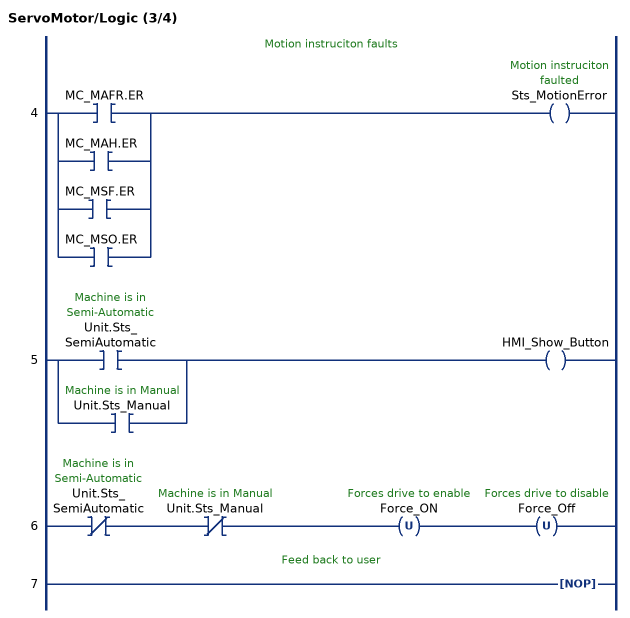
   // Motion instruciton faults
   4: [XIC(MC_MAFR.ER) ,XIC(MC_MAH.ER) ,XIC(MC_MSF.ER) ,XIC(MC_MSO.ER) ]OTE(Sts_MotionError);
   5: [XIC(Unit.Sts_SemiAutomatic) ,XIC(Unit.Sts_Manual) ]OTE(HMI_Show_Button);
   6: XIO(Unit.Sts_SemiAutomatic)XIO(Unit.Sts_Manual)OTU(Force_ON)OTU(Force_Off);
   // Feed back to user
   7: NOP();
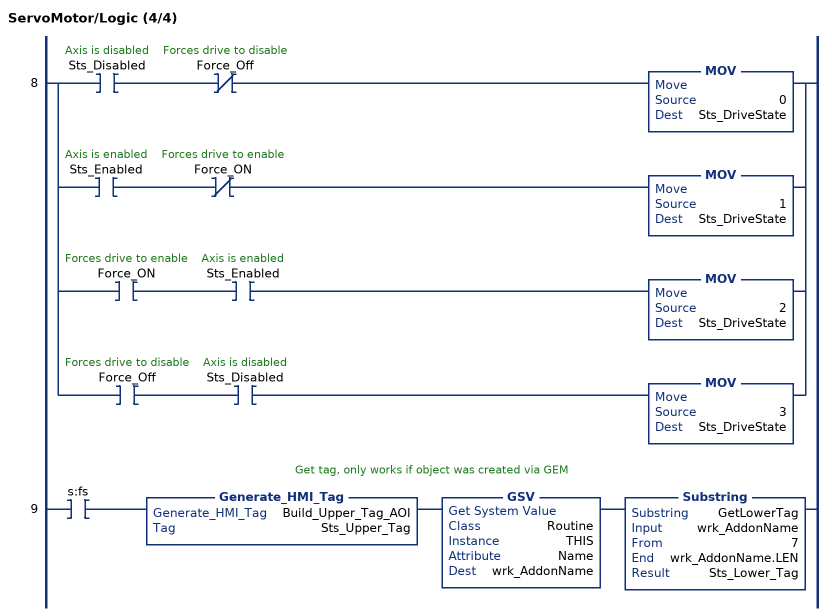
   8: [XIC(Sts_Disabled) XIO(Force_Off) MOV(0,Sts_DriveState) ,XIC(Sts_Enabled) XIO(Force_ON) MOV(1,Sts_DriveState) ,XIC(Force_ON) XIC(Sts_Enabled) MOV(2,Sts_DriveState) ,XIC(Force_Off) XIC(Sts_Disabled) MOV(3,Sts_DriveState) ];
   // Get tag, only works if object was created via GEM
   9: XIC(s:fs)Generate_HMI_Tag(Build_Upper_Tag_AOI,Sts_Upper_Tag)GSV(Routine,THIS,Name,wrk_AddonName)Substring(GetLowerTag,wrk_AddonName,7,wrk_AddonName.LEN,Sts_Lower_Tag);
END_ROUTINE

ROUTINE Prescan   (* structured text *)
   ////////////////////////////////////////////////////////////
   //   Copyright (c)
   //------------------------------------------------------------
   //   Routine: Prescan
   //   Author: WPI\tom.reit
   //   Created: 18-1-2023
   //------------------------------------------------------------
   //   Description:
   //
   //
   //   History:
   //
   ////////////////////////////////////////////////////////////
   MC_MAH.FLAGS		:=0;
   MC_MAFR.FLAGS		:=0;
   MC_MSF.FLAGS		:=0;
   MC_MSO.FLAGS		:=0;
   
END_ROUTINE
END_ADD_ON_INSTRUCTION

ADD_ON_INSTRUCTION SimpleDrive_Digital   (* revision 1.0 *)
VAR_OUTPUT
   O_Start : BOOL; {required}   // Phyical output to start drive
END_VAR
VAR_INPUT
   Start : BOOL; {visible}   // Starts the drive
   I_Fault : BOOL; {visible}   // Fault input
END_VAR
VAR_OUTPUT
   Sts_Faulted : BOOL; {visible}   // Drive Faulted
   Sts_Drive_Running : BOOL; {visible}   // Motor is running
END_VAR
VAR_INPUT
   Force_ON : BOOL; {visible}   // Forces the drive on
   Force_Off : BOOL; {visible}   // Forces the drive off
END_VAR
VAR_OUTPUT
   Sts_DriveState : DINT; {visible}   // Drive states for HMI 0=Drive not active 1=Drive active 2=Manual turned on 3=Manual turned off
   HMI_Show_Button : BOOL;   // only for HMI control
END_VAR
VAR_IN_OUT
   Unit : ISA_TR_88_00_02; {required}
END_VAR
VAR
   Sts_Upper_Tag : STRING; {access Read Only}   // Unit_EM
   Sts_Lower_Tag : STRING; {access Read Only}   // Object Name
   GetLowerTag : Substring; {access None}
   Build_Upper_Tag_AOI : Generate_HMI_Tag; {access None}
   wrk_AddonName : STRING; {access None}
   T_Decel : TIMER := (PRE := 5000); {access None}
END_VAR

ROUTINE Logic   (* ladder *)
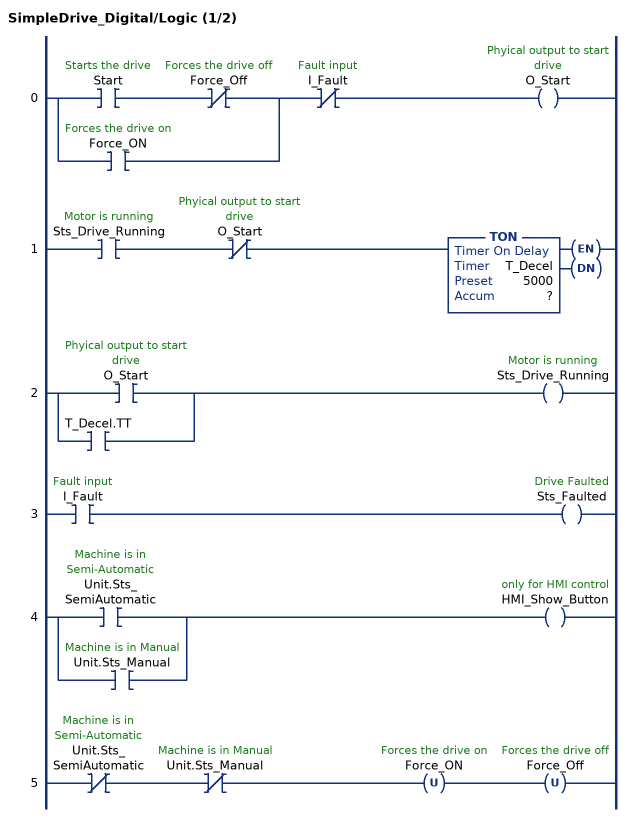
   0: [XIC(Start) XIO(Force_Off) ,XIC(Force_ON) ]XIO(I_Fault)OTE(O_Start);
   1: XIC(Sts_Drive_Running)XIO(O_Start)TON(T_Decel,?,?);
   2: [XIC(O_Start) ,XIC(T_Decel.TT) ]OTE(Sts_Drive_Running);
   3: XIC(I_Fault)OTE(Sts_Faulted);
   4: [XIC(Unit.Sts_SemiAutomatic) ,XIC(Unit.Sts_Manual) ]OTE(HMI_Show_Button);
   5: XIO(Unit.Sts_SemiAutomatic)XIO(Unit.Sts_Manual)OTU(Force_ON)OTU(Force_Off);
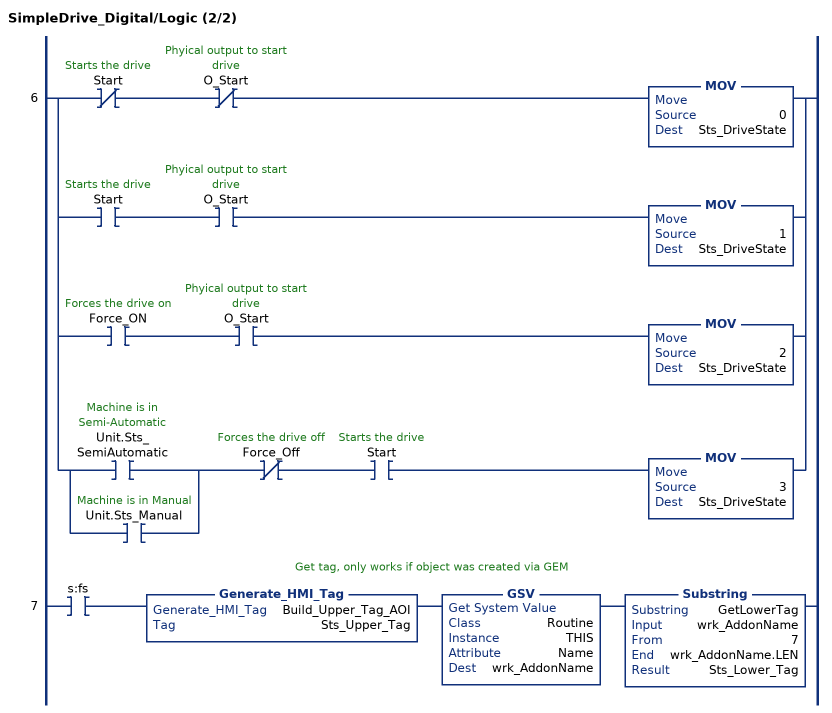
   6: [XIO(Start) XIO(O_Start) MOV(0,Sts_DriveState) ,XIC(Start) XIC(O_Start) MOV(1,Sts_DriveState) ,XIC(Force_ON) XIC(O_Start) MOV(2,Sts_DriveState) ,[XIC(Unit.Sts_SemiAutomatic) ,XIC(Unit.Sts_Manual) ] XIO(Force_Off) XIC(Start) MOV(3,Sts_DriveState) ];
   // Get tag, only works if object was created via GEM
   7: XIC(s:fs)Generate_HMI_Tag(Build_Upper_Tag_AOI,Sts_Upper_Tag)GSV(Routine,THIS,Name,wrk_AddonName)Substring(GetLowerTag,wrk_AddonName,7,wrk_AddonName.LEN,Sts_Lower_Tag);
END_ROUTINE
END_ADD_ON_INSTRUCTION

ADD_ON_INSTRUCTION SimpleDrive_SpeedControl   (* revision 1.0 *)
VAR_IN_OUT
   Unit : ISA_TR_88_00_02; {required}
END_VAR
VAR_INPUT
   cnf_Min_Speed : REAL; {visible}   // Min speed the drive may run at
   cnf_Max_Speed : REAL; {visible}   // Max speed the drive may run at
   Speed : REAL; {visible}   // Requested speed
   Start : BOOL; {visible}   // Starts the drive
   Force_ON : BOOL; {visible}   // Forces the drive on
   Force_Off : BOOL; {visible}   // Forces the drive off
END_VAR
VAR_OUTPUT
   O_Start : BOOL; {required}   // Phyical output to start drive
   O_Speed : REAL; {required}   // Output speed
END_VAR
VAR_INPUT
   I_Fault : BOOL; {visible}   // Fault input
END_VAR
VAR_OUTPUT
   Sts_Faulted : BOOL; {visible}   // Drive Faulted
   Sts_Drive_Running : BOOL; {visible}   // Motor is running
   Sts_DriveState : DINT;   // Drive states for HMI 0=Drive not active 1=Drive active 2=Manual turned on 3=Manual turned off
   HMI_Show_Button : BOOL;   // only for HMI control
END_VAR
VAR
   Sts_Upper_Tag : STRING; {access Read Only}   // Unit_EM
   Sts_Lower_Tag : STRING; {access Read Only}   // Object Name
   GetLowerTag : Substring; {access None}
   Build_Upper_Tag_AOI : Generate_HMI_Tag; {access None}
   wrk_AddonName : STRING; {access None}
   SpeedDrive : AnalogOutput; {access None}
   T_Decel : TIMER := (PRE := 5000); {access None}
END_VAR

ROUTINE Logic   (* ladder *)
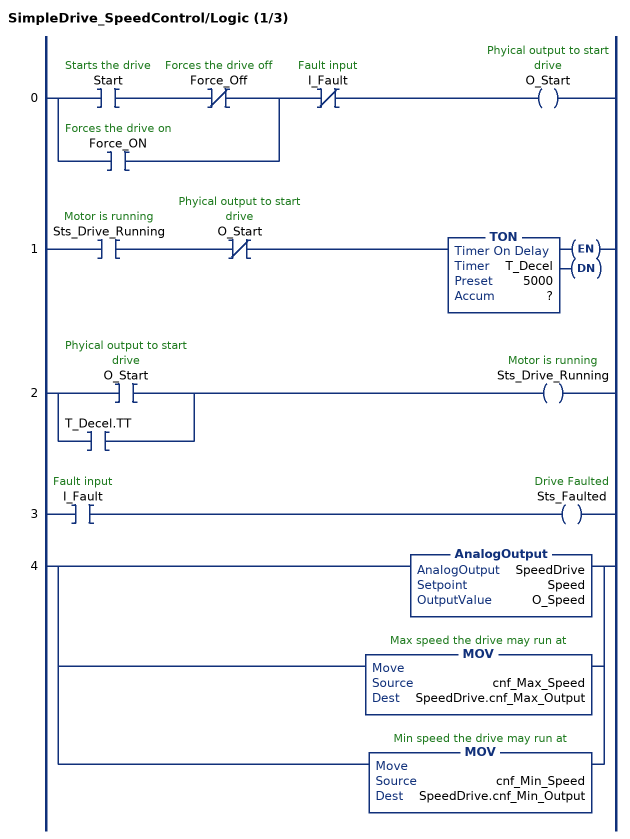
   0: [XIC(Start) XIO(Force_Off) ,XIC(Force_ON) ]XIO(I_Fault)OTE(O_Start);
   1: XIC(Sts_Drive_Running)XIO(O_Start)TON(T_Decel,?,?);
   2: [XIC(O_Start) ,XIC(T_Decel.TT) ]OTE(Sts_Drive_Running);
   3: XIC(I_Fault)OTE(Sts_Faulted);
   4: [AnalogOutput(SpeedDrive,Speed,O_Speed) ,MOV(cnf_Max_Speed,SpeedDrive.cnf_Max_Output) ,MOV(cnf_Min_Speed,SpeedDrive.cnf_Min_Output) ];
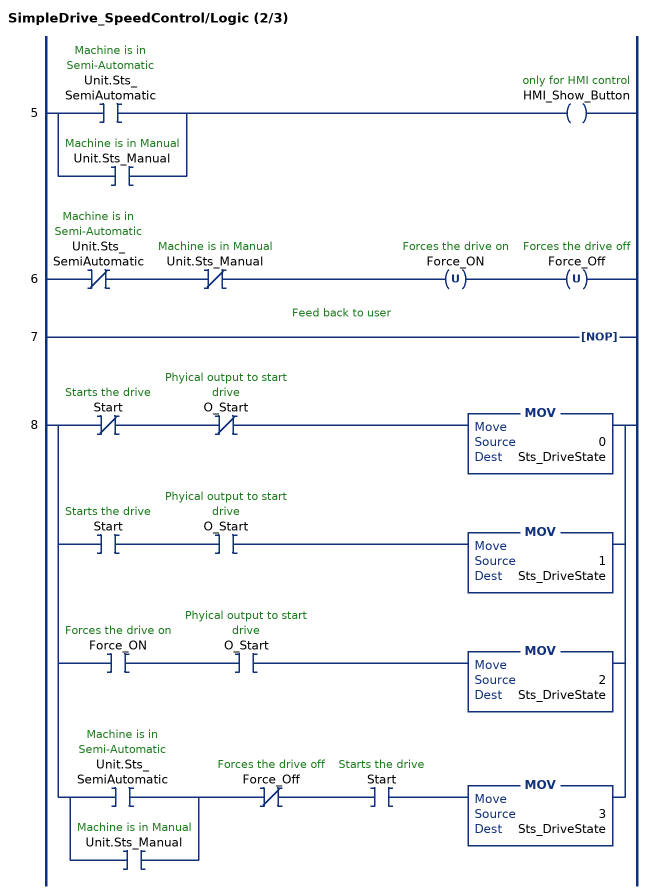
   5: [XIC(Unit.Sts_SemiAutomatic) ,XIC(Unit.Sts_Manual) ]OTE(HMI_Show_Button);
   6: XIO(Unit.Sts_SemiAutomatic)XIO(Unit.Sts_Manual)OTU(Force_ON)OTU(Force_Off);
   // Feed back to user
   7: NOP();
   8: [XIO(Start) XIO(O_Start) MOV(0,Sts_DriveState) ,XIC(Start) XIC(O_Start) MOV(1,Sts_DriveState) ,XIC(Force_ON) XIC(O_Start) MOV(2,Sts_DriveState) ,[XIC(Unit.Sts_SemiAutomatic) ,XIC(Unit.Sts_Manual) ] XIO(Force_Off) XIC(Start) MOV(3,Sts_DriveState) ];
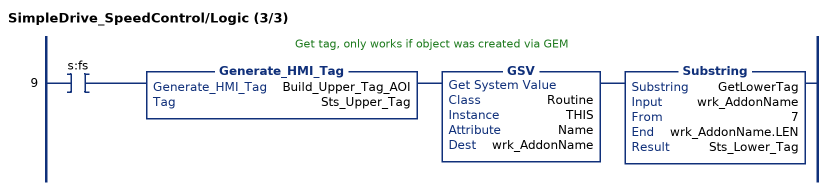
   // Get tag, only works if object was created via GEM
   9: XIC(s:fs)Generate_HMI_Tag(Build_Upper_Tag_AOI,Sts_Upper_Tag)GSV(Routine,THIS,Name,wrk_AddonName)Substring(GetLowerTag,wrk_AddonName,7,wrk_AddonName.LEN,Sts_Lower_Tag);
END_ROUTINE
END_ADD_ON_INSTRUCTION

ADD_ON_INSTRUCTION Substring   (* revision 1.0, vendor WPI *)
VAR_IN_OUT
   Input : STRING; {required}   // String to substring
END_VAR
VAR_INPUT
   From : INT; {required}   // where to start substringing
   End : DINT; {required}   // Where to end the substring
END_VAR
VAR_IN_OUT
   Result : STRING; {required}   // Result from substring
END_VAR
VAR
   i : DINT; {access None}   // local index
END_VAR

ROUTINE Logic   (* structured text *)
   #region Prevent controler fault
   		if From >= 80 	then From	:=80;	end_if;		// starting pos can never be higher then 80
   		if -1 	>= From then From	:=0; 	end_if;		// starting pos can never be lower then 0
   
   		if End >= 81 	then From	:=81;	end_if;		// ending pos can never be higher then 81
   		if -1 	>= End 	then End	:=1; 	end_if;		// ending pos can never be lower then 1
   	if From >= End then
   		End						:=	From+1;				// if end is lower or equal to from, no boundries are set for a substring. to prevent this add 1 to end to substring only 1 char.
   	end_if;
   #endregion
   #region Substring
   	#region clear previous data
   		for i := 0 to 81 do
   			Result.DATA[i] 		:=	0;					// set all data back to 0
   		end_for;
   		Result.LEN				:=	0;					// string length is set back to 0
   	#endregion
   	for i := From to End do
   		Result.DATA[i-From]		:=	Input.DATA[i];		// add substring data to Result, shift Index to start from Result.data[0] -> Result.data[1] -> Result.data[2] etc.
   	end_for;
   	Result.LEN					:=	End-From;			// set string length
   #endregion
END_ROUTINE
END_ADD_ON_INSTRUCTION

ADD_ON_INSTRUCTION Valve_V2   (* revision 1.0, ExecutePrescan *)
VAR_IN_OUT
   PackML : ISA_TR_88_00_02; {required}
END_VAR
VAR_INPUT
   Turn_On : BOOL := 1; {visible}   // Turn on the valve by program
END_VAR
VAR_OUTPUT
   Valve_Out : BOOL; {access Read Only, required}   // Connection to valve tag
END_VAR
VAR_INPUT
   Reset : BOOL; {visible}   // Reset valve timers
   cnf_NO_or_NC : BOOL; {visible}   // normally open or normally closed 0 = NO 1 = NC
   cnf_Retain_By_Fault : BOOL := 1; {visible}   // if the machine faulted, while the valve was open. it stays open.
   cnf_Feedback : BOOL := 1; {visible}   // set to true if valve has feedback
   Feedback_signal : BOOL; {required}   // feedback signal from valve if valve has no feedback use Valve_Out tag
END_VAR
VAR_OUTPUT
   HMI_color : DINT; {access Read Only}   // color of valve
   Sts_Faulted : BOOL; {access Read Only, visible}   // Valve did not open within feedback time
   Sts_Valve_open : BOOL; {access Read Only, visible}   // valve is open according to feedback
   Sts_Valve_Closed : BOOL; {access Read Only, visible}   // valve is closed according to feedback
   Sts_Valve_Status : DINT; {access Read Only}   // indicator dint for HMI about valve state
   Sts_RetainedByFault : BOOL; {access Read Only, visible}   // Machine faulted, holding valve open or closed respectively
END_VAR
VAR_INPUT
   Force_Open : BOOL; {visible}   // Manual & Semiautomatic Forces valve to open
   Force_Closed : BOOL; {visible}   // Manual & Semiautomatic Forces valve to close
END_VAR
VAR_OUTPUT
   Sts_Show_HMIControls : BOOL;   // 0 = dont show 1 = Show controls
   HMI_Show_Button : BOOL; {access Read Only}   // allow HMI to press manual control button
END_VAR
VAR
   T_Switch_Time : TIMER[2] := ([0].PRE := 250, [1].PRE := 250); {access None}   // timer for valve to move from open to close or the otherway around
   wrk_hold_state : BOOL := 1; {access None}   // machine faulted, holding valve in current state until machine is resetted.
   ons_reset : BOOL; {access None}   // prevent continious reset
   T_Mem_Valve : TIMER[2] := ([0].PRE := 50, [1].PRE := 50); {access None}
   Wrk_Valve_Out : BOOL; {access None}   // local mem for retain by fault
   Manual_Turn_on : BOOL; {access None}   // local valve control
   wrk_AddonName : STRING := 'CM_002_CV01'; {access None}
   Sts_Upper_Tag : STRING; {access Read Only}   // Unit_EM
   Build_Upper_Tag_AOI : Generate_HMI_Tag; {access None}
   Sts_Lower_Tag : STRING; {access Read Only}   // Object Name
   GetLowerTag : Substring; {access None}
END_VAR

ROUTINE Logic   (* ladder *)
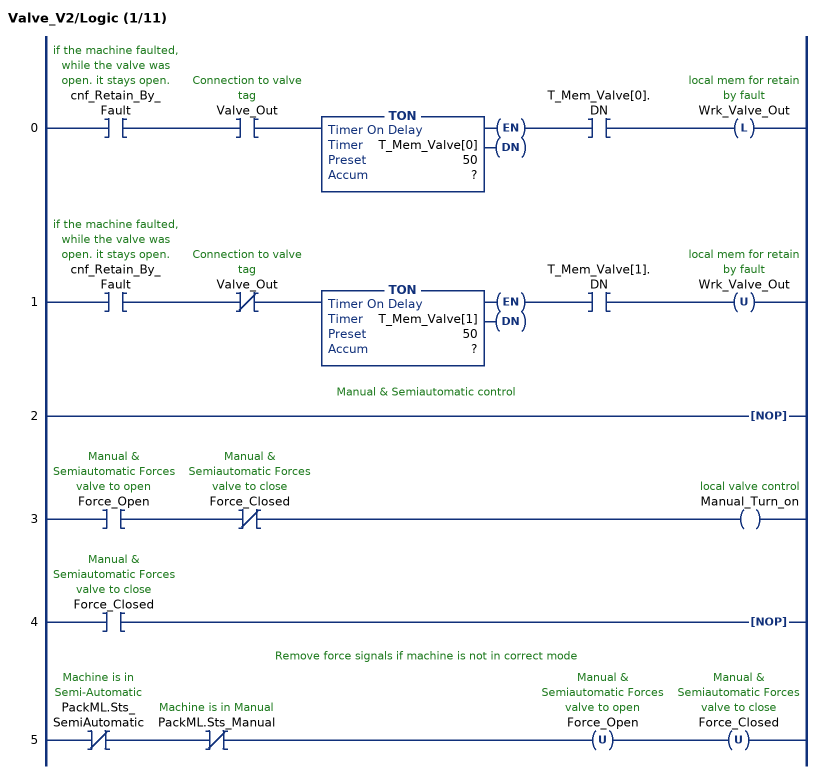
   0: XIC(cnf_Retain_By_Fault)XIC(Valve_Out)TON(T_Mem_Valve[0],?,?)XIC(T_Mem_Valve[0].DN)OTL(Wrk_Valve_Out);
   1: XIC(cnf_Retain_By_Fault)XIO(Valve_Out)TON(T_Mem_Valve[1],?,?)XIC(T_Mem_Valve[1].DN)OTU(Wrk_Valve_Out);
   // Manual & Semiautomatic control
   2: NOP();
   3: XIC(Force_Open)XIO(Force_Closed)OTE(Manual_Turn_on);
   4: XIC(Force_Closed)NOP();
   // Remove force signals if machine is not in correct mode
   5: XIO(PackML.Sts_SemiAutomatic)XIO(PackML.Sts_Manual)OTU(Force_Open)OTU(Force_Closed);
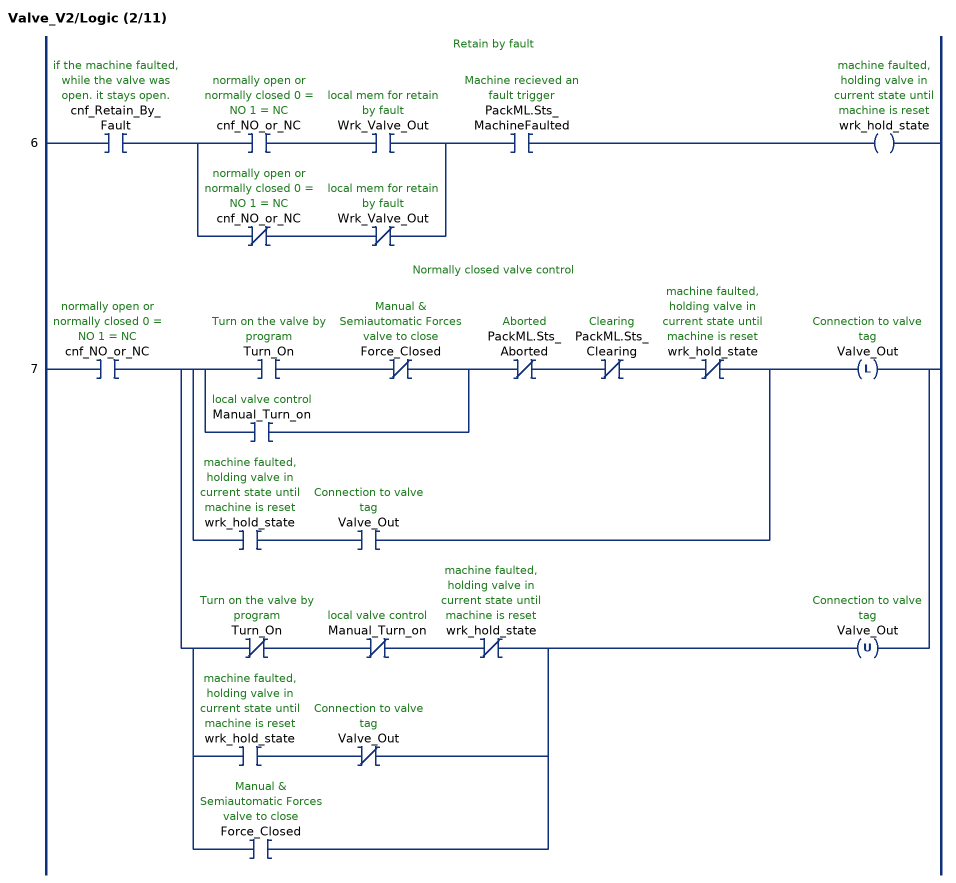
   // Retain by fault
   6: XIC(cnf_Retain_By_Fault)[XIC(cnf_NO_or_NC) XIC(Wrk_Valve_Out) ,XIO(cnf_NO_or_NC) XIO(Wrk_Valve_Out) ]XIC(PackML.Sts_MachineFaulted)OTE(wrk_hold_state);
   // Normally closed valve control
   7: XIC(cnf_NO_or_NC)[[[XIC(Turn_On) XIO(Force_Closed) ,XIC(Manual_Turn_on) ] XIO(PackML.Sts_Aborted) XIO(PackML.Sts_Clearing) XIO(wrk_hold_state) ,XIC(wrk_hold_state) XIC(Valve_Out) ] OTL(Valve_Out) ,[XIO(Turn_On) XIO(Manual_Turn_on) XIO(wrk_hold_state) ,XIC(wrk_hold_state) XIO(Valve_Out) ,XIC(Force_Closed) ] OTU(Valve_Out) ];
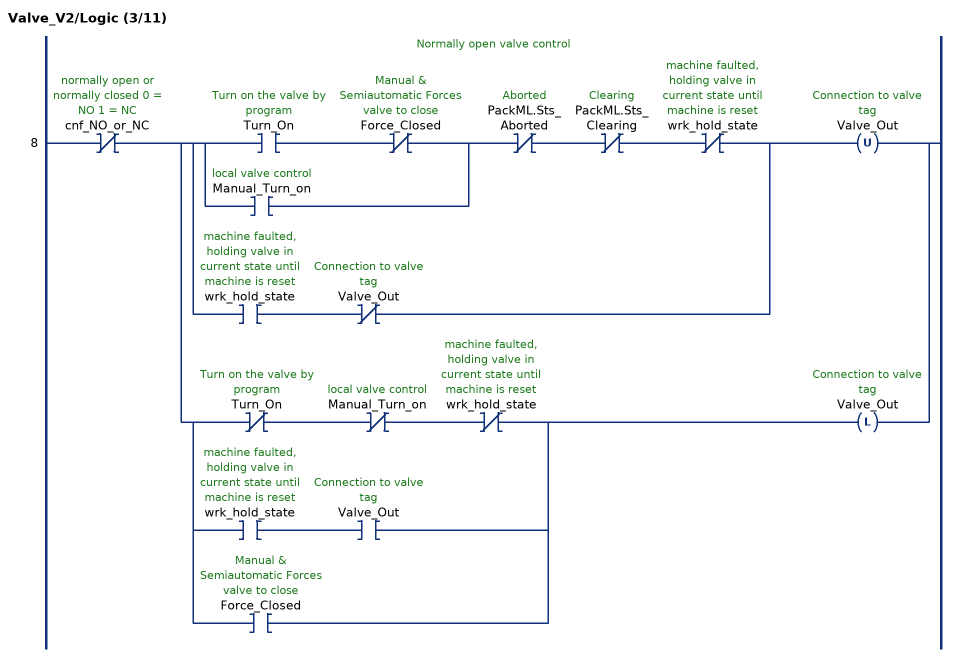
   // Normally open valve control
   8: XIO(cnf_NO_or_NC)[[[XIC(Turn_On) XIO(Force_Closed) ,XIC(Manual_Turn_on) ] XIO(PackML.Sts_Aborted) XIO(PackML.Sts_Clearing) XIO(wrk_hold_state) ,XIC(wrk_hold_state) XIO(Valve_Out) ] OTU(Valve_Out) ,[XIO(Turn_On) XIO(Manual_Turn_on) XIO(wrk_hold_state) ,XIC(wrk_hold_state) XIC(Valve_Out) ,XIC(Force_Closed) ] OTL(Valve_Out) ];
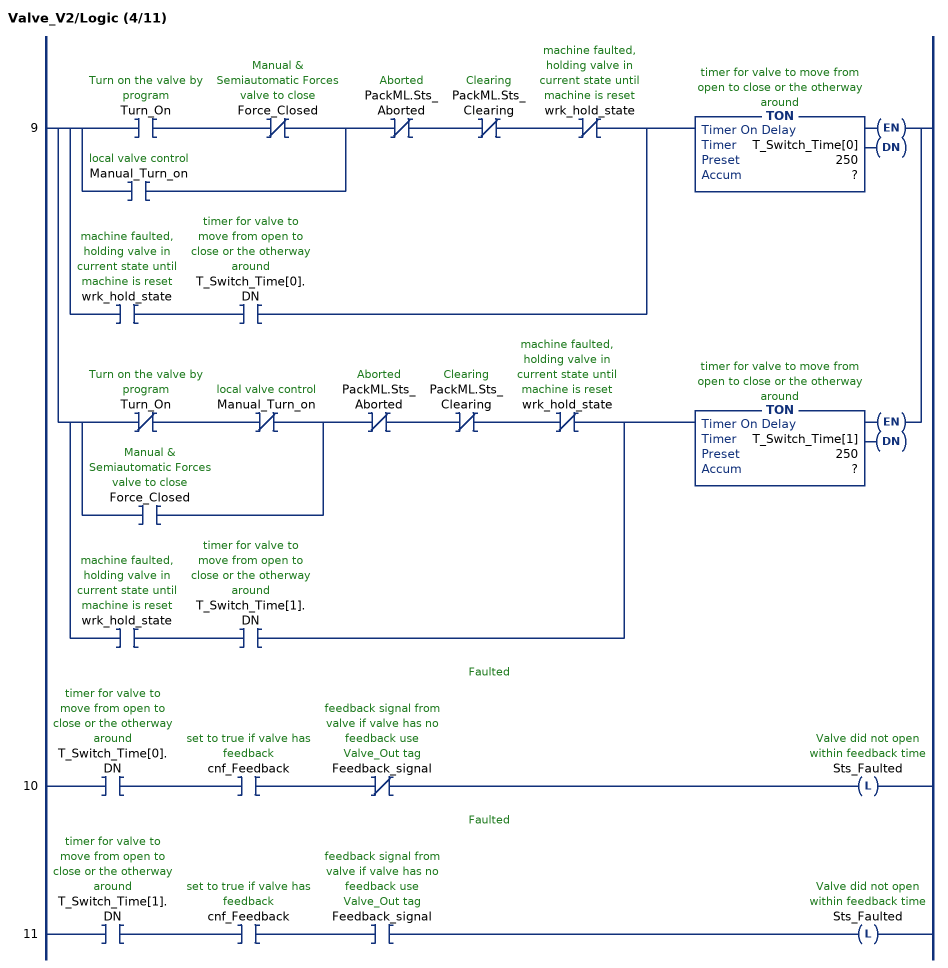
   9: [[[XIC(Turn_On) XIO(Force_Closed) ,XIC(Manual_Turn_on) ] XIO(PackML.Sts_Aborted) XIO(PackML.Sts_Clearing) XIO(wrk_hold_state) ,XIC(wrk_hold_state) XIC(T_Switch_Time[0].DN) ] TON(T_Switch_Time[0],?,?) ,[[XIO(Turn_On) XIO(Manual_Turn_on) ,XIC(Force_Closed) ] XIO(PackML.Sts_Aborted) XIO(PackML.Sts_Clearing) XIO(wrk_hold_state) ,XIC(wrk_hold_state) XIC(T_Switch_Time[1].DN) ] TON(T_Switch_Time[1],?,?) ];
   // Faulted
   10: XIC(T_Switch_Time[0].DN)XIC(cnf_Feedback)XIO(Feedback_signal)OTL(Sts_Faulted);
   // Faulted
   11: XIC(T_Switch_Time[1].DN)XIC(cnf_Feedback)XIC(Feedback_signal)OTL(Sts_Faulted);
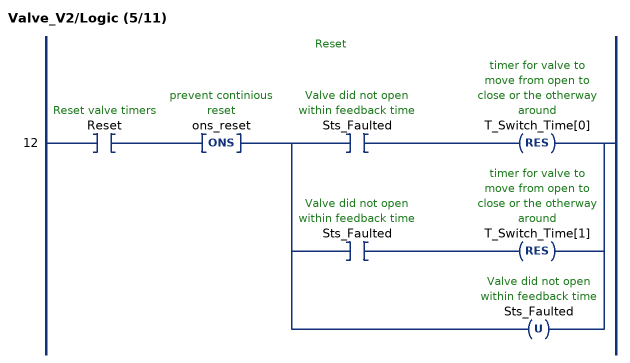
   // Reset
   12: XIC(Reset)ONS(ons_reset)[XIC(Sts_Faulted) RES(T_Switch_Time[0]) ,XIC(Sts_Faulted) RES(T_Switch_Time[1]) ,OTU(Sts_Faulted) ];
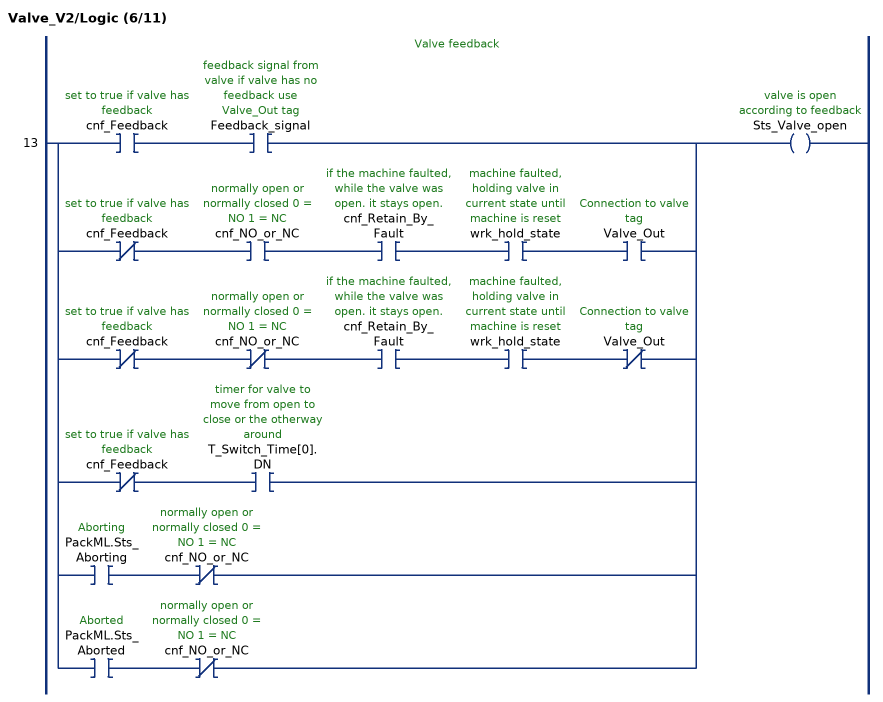
   // Valve feedback
   13: [XIC(cnf_Feedback) XIC(Feedback_signal) ,XIO(cnf_Feedback) XIC(cnf_NO_or_NC) XIC(cnf_Retain_By_Fault) XIC(wrk_hold_state) XIC(Valve_Out) ,XIO(cnf_Feedback) XIO(cnf_NO_or_NC) XIC(cnf_Retain_By_Fault) XIC(wrk_hold_state) XIO(Valve_Out) ,XIO(cnf_Feedback) XIC(T_Switch_Time[0].DN) ,XIC(PackML.Sts_Aborting) XIO(cnf_NO_or_NC) ,XIC(PackML.Sts_Aborted) XIO(cnf_NO_or_NC) ]OTE(Sts_Valve_open);
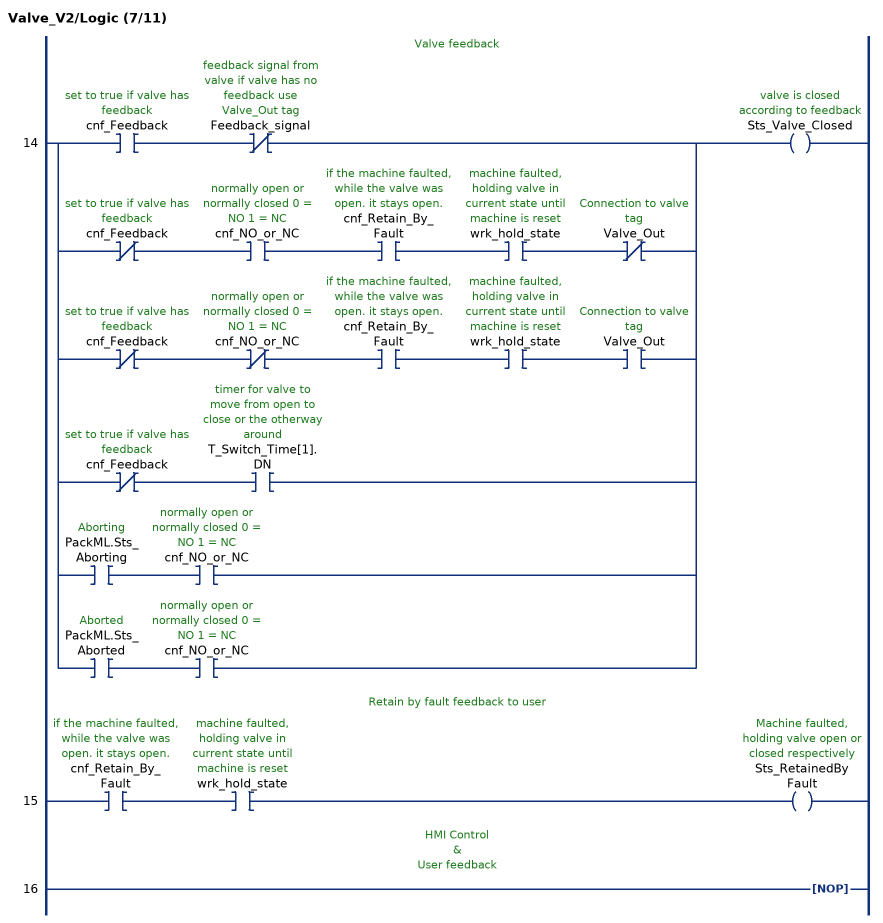
   // Valve feedback
   14: [XIC(cnf_Feedback) XIO(Feedback_signal) ,XIO(cnf_Feedback) XIC(cnf_NO_or_NC) XIC(cnf_Retain_By_Fault) XIC(wrk_hold_state) XIO(Valve_Out) ,XIO(cnf_Feedback) XIO(cnf_NO_or_NC) XIC(cnf_Retain_By_Fault) XIC(wrk_hold_state) XIC(Valve_Out) ,XIO(cnf_Feedback) XIC(T_Switch_Time[1].DN) ,XIC(PackML.Sts_Aborting) XIC(cnf_NO_or_NC) ,XIC(PackML.Sts_Aborted) XIC(cnf_NO_or_NC) ]OTE(Sts_Valve_Closed);
   // Retain by fault feedback to user
   15: XIC(cnf_Retain_By_Fault)XIC(wrk_hold_state)OTE(Sts_RetainedByFault);
   // HMI Control
   // &
   // User feedback
   16: NOP();
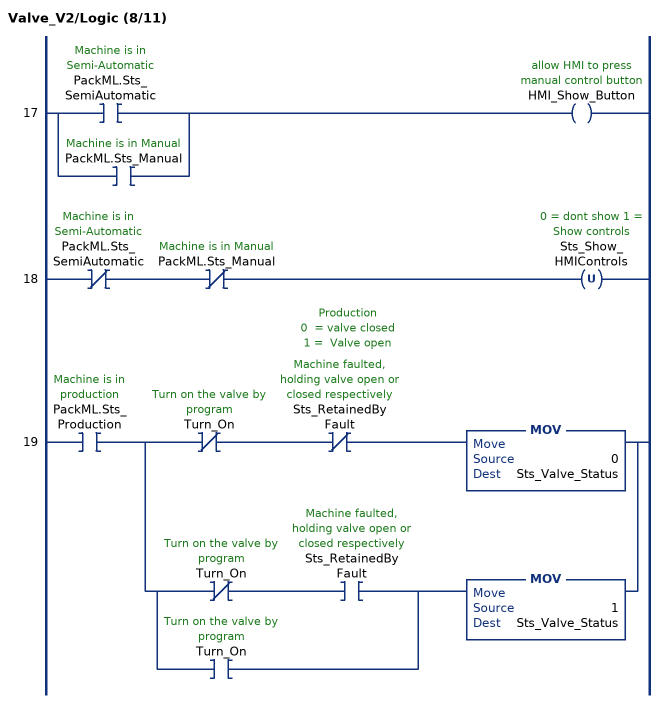
   17: [XIC(PackML.Sts_SemiAutomatic) ,XIC(PackML.Sts_Manual) ]OTE(HMI_Show_Button);
   18: XIO(PackML.Sts_SemiAutomatic)XIO(PackML.Sts_Manual)OTU(Sts_Show_HMIControls);
   // Production
   // 0  = valve closed
   // 1 =  Valve open
   19: XIC(PackML.Sts_Production)[XIO(Turn_On) XIO(Sts_RetainedByFault) MOV(0,Sts_Valve_Status) ,[XIO(Turn_On) XIC(Sts_RetainedByFault) ,XIC(Turn_On) ] MOV(1,Sts_Valve_Status) ];
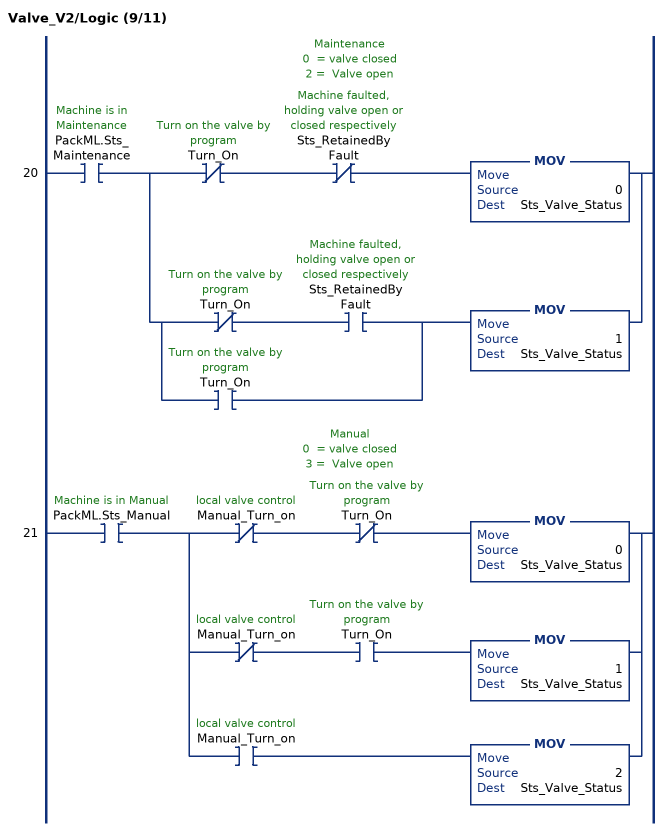
   // Maintenance
   // 0  = valve closed
   // 2 =  Valve open
   20: XIC(PackML.Sts_Maintenance)[XIO(Turn_On) XIO(Sts_RetainedByFault) MOV(0,Sts_Valve_Status) ,[XIO(Turn_On) XIC(Sts_RetainedByFault) ,XIC(Turn_On) ] MOV(1,Sts_Valve_Status) ];
   // Manual
   // 0  = valve closed
   // 3 =  Valve open
   21: XIC(PackML.Sts_Manual)[XIO(Manual_Turn_on) XIO(Turn_On) MOV(0,Sts_Valve_Status) ,XIO(Manual_Turn_on) XIC(Turn_On) MOV(1,Sts_Valve_Status) ,XIC(Manual_Turn_on) MOV(2,Sts_Valve_Status) ];
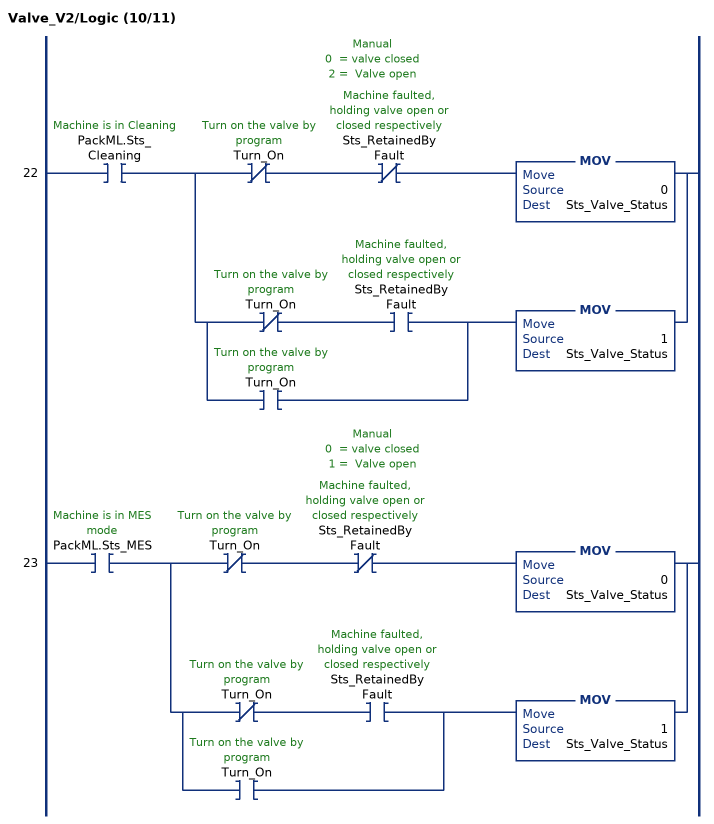
   // Manual
   // 0  = valve closed
   // 2 =  Valve open
   22: XIC(PackML.Sts_Cleaning)[XIO(Turn_On) XIO(Sts_RetainedByFault) MOV(0,Sts_Valve_Status) ,[XIO(Turn_On) XIC(Sts_RetainedByFault) ,XIC(Turn_On) ] MOV(1,Sts_Valve_Status) ];
   // Manual
   // 0  = valve closed
   // 1 =  Valve open
   23: XIC(PackML.Sts_MES)[XIO(Turn_On) XIO(Sts_RetainedByFault) MOV(0,Sts_Valve_Status) ,[XIO(Turn_On) XIC(Sts_RetainedByFault) ,XIC(Turn_On) ] MOV(1,Sts_Valve_Status) ];
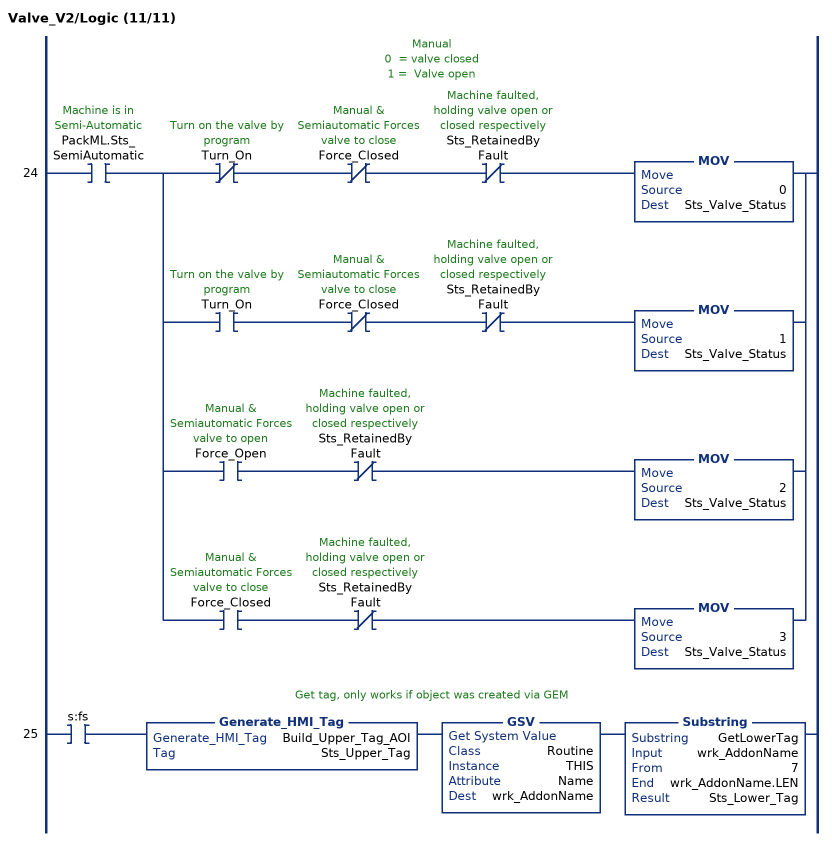
   // Manual
   // 0  = valve closed
   // 1 =  Valve open
   24: XIC(PackML.Sts_SemiAutomatic)[XIO(Turn_On) XIO(Force_Closed) XIO(Sts_RetainedByFault) MOV(0,Sts_Valve_Status) ,XIC(Turn_On) XIO(Force_Closed) XIO(Sts_RetainedByFault) MOV(1,Sts_Valve_Status) ,XIC(Force_Open) XIO(Sts_RetainedByFault) MOV(2,Sts_Valve_Status) ,XIC(Force_Closed) XIO(Sts_RetainedByFault) MOV(3,Sts_Valve_Status) ];
   // Get tag, only works if object was created via GEM
   25: XIC(s:fs)Generate_HMI_Tag(Build_Upper_Tag_AOI,Sts_Upper_Tag)GSV(Routine,THIS,Name,wrk_AddonName)Substring(GetLowerTag,wrk_AddonName,7,wrk_AddonName.LEN,Sts_Lower_Tag);
END_ROUTINE
